// TIA Portal project "CLU" (V13)

(* hardware
DEVICE "S7-1200 station_1"  S7-1200 Station
   slot 0: "Telaio di montaggio_0"  Rack  V1.0
   slot 1: "S7_1200"  CPU 1214C DC/DC/DC  6ES7 214-1AG40-0XB0  V4.1
   slot 2: "DI 8/DQ 8x24VDC_1"  6ES7 223-1BH32-0XB0  V2.0
   slot 3: "DI 16/DQ 16x24VDC_1"  6ES7 223-1BL32-0XB0  V2.0
   slot 3: "Scheda di batteria_1"  6ES7 297-0AX30-0XA0  V1.0
   slot 4: "AI 8x13BIT_1"  6ES7 231-4HF32-0XB0  V2.0
   slot 5: "AI 8x13BIT_2"  6ES7 231-4HF32-0XB0  V2.0
   slot 6: "AQ 4x14BIT_1"  6ES7 232-4HD32-0XB0  V2.0
   slot 101: "CM 1241 (RS422/485)_1"  6ES7 241-1CH32-0XB0  V2.0
DEVICE "DISPLAY_KTP400"  KTP400 Basic color PN
   slot 0: "HMI"  HMI  6AV6 647-0AK11-3AX0  12.0.0.0
   slot 1: "HMI_RT_1"  KTP400 Basic color PN  6AV6 647-0AK11-3AX0  12.0.0.0
   slot 5: "DISPLAY_KTP400.IE_CP_1"  Interfaccia PROFINET
      slot 1: "PROFINET Interface_1"  Interfaccia PROFINET
         slot 1: "Porta_2"  Porta
*)

// ===== PLC "S7_1200"  CPU 1214C DC/DC/DC =====

VAR_GLOBAL   // PLC tag table "Tabella delle variabili standard"
   "ATTIVA_PRG" AT %M2.0 : Bool;   // Attiva il programma principale
   "System_Byte" AT %MB0 : Byte;
   "FirstScan" AT %M0.0 : Bool;   // Contatto chiuso solo alla prima scansiona
   "DiagStatusUpdate" AT %M0.1 : Bool;
   "AlwaysTRUE" AT %M0.2 : Bool;   // Contatto sempre chiuso
   "AlwaysFALSE" AT %M0.3 : Bool;   // Contatto sempre aperto
   "Clock_1.25Hz" AT %M1.4 : Bool;
   "Clock_1Hz" AT %M1.5 : Bool;
   "Clock_0.625Hz" AT %M1.6 : Bool;
   "Clock_0.5Hz" AT %M1.7 : Bool;
   "tasto_REMOTO" AT %I0.1 : Bool;
   "tasto_OFF" AT %I0.2 : Bool;
   "tasto_ON" AT %I0.3 : Bool;
   "tasto_ANODICA" AT %I0.4 : Bool;
   "tasto_RESET" AT %I0.5 : Bool;
   "led_LOCALE" AT %Q0.0 : Bool;
   "led_REMOTO" AT %Q0.1 : Bool;
   "led_OFF" AT %Q0.2 : Bool;
   "led_ON" AT %Q0.3 : Bool;
   "led_ANODICA" AT %Q0.4 : Bool;
   "led_RESET" AT %Q0.5 : Bool;
   "in_FLUSSO_LQD_TUBO_SEGNALE" AT %I0.6 : Bool;
   "in_FLUSSO_LQD_SS_SEGNALE" AT %I0.7 : Bool;
   "in_MAX_TEMP_LQD_SS_OK" AT %I1.0 : Bool;
   "in_MIN_PRESSIONE_LQD_SS_OK" AT %I1.1 : Bool;
   "in_INTERLOCK_OK" AT %I1.3 : Bool;
   "in_FLUSSO_LQD_TUBO_OK" AT %I1.4 : Bool;
   "in_FLUSSO_LQD_SS_OK" AT %I1.5 : Bool;
   "in_MAX_IG2_OK" AT %I2.0 : Bool;
   "adc_FWD_TUBO" AT %IW5 : Word;
   "adc_RFL_TUBO" AT %IW7 : Word;
   "adc_TENSIONE_ANODICA" AT %IW21 : Word;
   "adc_CORRENTE_ANODICA" AT %IW23 : Word;
   "adc_TENSIONE_G1" AT %IW25 : Word;
   "adc_CORRENTE_G1" AT %IW27 : Word;
   "adc_TENSIONE_G2" AT %IW29 : Word;
   "adc_CORRENTE_G2" AT %IW31 : Word;
   "led_RIFLESSA" AT %Q0.6 : Bool;
   "led_TEMPERTURA" AT %Q0.7 : Bool;
   "led_COOLING" AT %Q1.0 : Bool;
   "led_PREALLAME" AT %Q1.1 : Bool;
   "led_REDUCED" AT %Q2.0 : Bool;
   "led_NOMINAL" AT %Q2.1 : Bool;
   "in_PRESSIONE_ARIA_CAVITA_OK" AT %I3.0 : Bool;
   "in_PRESSIONE_ARIA_FILAMENTO_OK" AT %I3.1 : Bool;
   "in_ALIMENTAZIONE_G1_OK" AT %I3.3 : Bool;
   "in_ALIMENTAZIONE_G2_OK" AT %I3.4 : Bool;
   "in_MAX_TEMP_LQD_TUBO_OK" AT %I3.5 : Bool;
   "in_MIN_PRESSIONE_LQD_TUBO_OK" AT %I3.6 : Bool;
   "in_SLAVE_PREALLARME" AT %I2.7 : Bool;   // Ingresso modalità Master/Slave
   "in_CONDUCIMETRO_OK" AT %I4.0 : Bool;
   "in_ALTA_TENSIONE_OK" AT %I4.1 : Bool;
   "in_MAX_TEMP_TRASF_AT_OK" AT %I4.2 : Bool;
   "in_MANCANZA_FASE_OK" AT %I4.4 : Bool;
   "in_IGNITRON_OK" AT %I4.5 : Bool;
   "in_MAX_IA_OK" AT %I4.6 : Bool;
   "in_VALVOLA_CAVITA_OK" AT %I4.7 : Bool;
   "out_ON_PREAMPLIFICATORE" AT %Q4.6 : Bool;
   "out_ON_DRIVER" AT %Q4.7 : Bool;
   "out_ON_CW" AT %Q2.2 : Bool;
   "out_VENTILAZIONE_CAVITA" AT %Q3.0 : Bool;
   "out_SLAVE_RESET" AT %Q3.1 : Bool;   // Uscita modalità Master/Slave
   "out_ALIMENTAZIONE_FILAMENTO" AT %Q3.2 : Bool;
   "out_PARZIALIZZATORE_FILAMENTO" AT %Q4.4 : Bool;
   "out_ALIMENTAZIONE_G1" AT %Q3.3 : Bool;
   "out_PARZIALIZZATORE_AT" AT %Q4.5 : Bool;
   "out_ALIMENTAZIONE_G2" AT %Q3.4 : Bool;
   "out_G2" AT %Q3.5 : Bool;
   "adc_CORRENTE_FILAMENTO" AT %IW33 : Word;
   "adc_ANALOGICA_7" AT %IW35 : Word;   // DISPONIBILE ANALOGICA
   "tasto_LOCALE" AT %I0.0 : Bool;
   "out_SLAVE_ON" AT %Q2.3 : Bool;   // Uscita modalità Master/Slave
   "in_COAX_POS_B" AT %I1.2 : Bool;
   "in_COAX_POS_A" AT %I2.1 : Bool;
   "in_SAFETY_MODULE_OK" AT %I4.3 : Bool;
   "out_COAX" AT %Q2.4 : Bool;   // Comando posizione Coassiale (S)=B, (R)=A
   "out_SLAVE_OFF" AT %Q2.5 : Bool;   // Uscita modalità Master/Slave
   "out_ON_AMP1" AT %Q3.6 : Bool;
   "out_ON_AMP2" AT %Q3.7 : Bool;
   "out_IGNITRON" AT %Q4.0 : Bool;
   "out_SLAVE_ALLARME" AT %Q4.2 : Bool;   // Uscita modalità Master/Slave
   "out_SLAVE_ANODICA_OFF" AT %Q4.1 : Bool;   // Uscita modalità Master/Slave
   "adc_TEMP_LQDin_SS" AT %IW11 : Word;
   "adc_TEMP_LQDout_SS" AT %IW13 : Word;
   "adc_TEMP_LQDout_Tubo" AT %IW15 : Word;
   "adc_TEMP_LQDin_Tubo" AT %IW17 : Word;
   "adc_FWD_SS" AT %IW9 : Word;
   "adc_RFL_SS" AT %IW19 : Word;
   "adc_ANALOGICA_1" AT %IW38 : Word;
   "adc_ANALOGICA_2" AT %IW40 : Word;
   "in_SLAVE_ON" AT %I2.2 : Bool;   // Ingresso modalità Master/Slave
   "in_SLAVE_OFF" AT %I2.3 : Bool;   // Ingresso modalità Master/Slave
   "in_SLAVE_ANODICA_ON" AT %I2.4 : Bool;   // Ingresso modalità Master/Slave
   "in_SLAVE_ANODICA_OFF" AT %I2.5 : Bool;   // Ingresso modalità Master/Slave
   "in_SLAVE_ALLARME" AT %I2.6 : Bool;   // Ingresso modalità Master/Slave
   "in_SELECT_MODE" AT %I3.2 : Bool;   // Ingresso modalità Master/Slave
   "out_SLAVE_ANODICA_ON" AT %Q2.6 : Bool;
   "out_SLAVE_PREALLARME" AT %Q4.3 : Bool;   // Uscita modalità Master/Slave
   "out_CW_PULSED_TRIGGER" AT %Q2.7 : Bool;
   "in_SLAVE_RESET" AT %I3.7 : Bool;   // Ingresso modalità Master/Slave
   "dac_out_VA" AT %QW5 : Word;   // Uscita analogica regolatore Tensione di anodica
   "dac_out_VG2" AT %QW7 : Word;   // Uscita analogica regolatore Tensione di anodica
   "dac_out_VG1" AT %QW9 : Word;   // Uscita analogica regolatore Tensione di anodica
   "dac_out_VF" AT %QW11 : Word;   // Uscita analogica regolatore Tensione di anodica
END_VAR

DATA_BLOCK "STATO"   // DB1
TITLE = STATO AMPLIFICATORE
{ S7_Optimized_Access := 'FALSE' }
AUTHOR : Dario
VERSION : 0.1
// Blocco dati dello stato generale dell'amplificatore.
   VAR RETAIN
      stato_LOCALE : Bool;
      stato_STANDBY : Bool;
      stato_ANODICA : Bool;
      stato_ALLARME : Bool;
      stato_BLOCCO : Bool;
      stato_MODO_PULSED : Bool;
      stato_MODO_CW : Bool;
      stato_SOLO_SS : Bool;
      stato_NORMALE : Bool;
      stato_MASTER : Bool;
      stato_SLAVE : Bool;
   END_VAR
   VAR
      stato_RFridotta : Bool;
      stato_RFnominale : Bool;
   END_VAR
   VAR RETAIN
      stato_sogliaROS_Tubo : Word;
      stato_sogliaROS400kW : Word;
      stato_sogliaROS_SS_Pulsed : Word;
      "stato sogliaROS_SS_CW" : Word;
      stato_AQNdelay : Word;
      stato_LimiterInputRF : Word;
      stato_sogliaRIDOTTA : Word;
   END_VAR
   VAR
      stato_sogliaNOMINALE : Word;
   END_VAR
   VAR RETAIN
      stato_RFtotaleParziale : Bool;
   END_VAR
   VAR
      stato_DISPLAY_1 : Word;
      stato_DISPLAY_2 : Word;
      stato_DISPLAY_3 : Word;
      stato_DISPLAY_4 : Word;
      stato_DISPLAY_5 : Word;
      stato_DISPLAY_6 : Word;
   END_VAR
   VAR RETAIN
      stato_AdjFWDTubo : Word;
      stato_AdjRFLTubo : Word;
      stato_AdjFWDSS : Word;
      stato_AdjRFLSS : Word;
      stato_AdjFWDTotale : Word;
      stato_AdjRFLTotale : Word;
   END_VAR
   VAR
      stato_Data : DTL;
   END_VAR
   VAR RETAIN
      stato_ADDR_1 : Byte;
      stato_ADDR_2 : Byte;
      stato_ADDR_3 : Byte;
      stato_ADDR_4 : Byte;
      stato_PORT : UInt;
      stato_ADJ_ANODICA_PULSED : Word;
      stato_ADJ_ANODICA_CW : Word;
      stato_VOLTAGGIO_G1 : DInt;
      stato_VOLTAGGIO_G2 : Word;
      stato_VOLTAGGIO_FILAMENTO : Word;
      stato_REGOLAZIONE_VG1 : Word;
      stato_adj_VA : Word;
      stato_adj_VG1 : Word;
      stato_adj_VG2 : Word;
      stato_adj_VF : Word;
      stato_ScaleVA : Word;
      stato_ScaleVG1 : Word;
      stato_ScaleVG2 : Word;
      stato_ScaleIF : Word;
      stato_ScaleIA : Word;
      stato_ScaleIG1 : Word;
      stato_ScaleIG2 : Word;
   END_VAR
   VAR
      allarme_FLUSSO_LQD_TUBO : Bool;
      allarme_FLUSSO_LQD_SS : Bool;
      allarme_PRESSIONE_MIN_LQD_TUBO : Bool;
      allarme_PRESSIONE_MAX_LQD_TUBO : Bool;
      allarme_PRESSIONE_LQD_SS : Bool;
      allarme_INTERLOCK_RF : Bool;
      allarme_INTERLOCK_GENERALE : Bool;
      allarme_CONDUCIMETRO : Bool;
      allarme_MAX_IA : Bool;
      allarme_MAX_IG1 : Bool;
      allarme_MAX_IG2 : Bool;
      allarme_MAX_IG2_SW : Bool;
      allarme_TEMPERATURA_LQD_TUBO : Bool;
      allarme_TEMPERATURA_LQD_SS : Bool;
      allarme_TEMPERATURA_LQD_DUMMY : Bool;
      allarme_TEMPERATURA_AT : Bool;
      allarme_IGNITRON : Bool;
      allarme_ROS_Tubo : Bool;
      allarme_ROS_SS : Bool;
      allarme_No_Aria_Cavità : Bool;
      allarme_ROS_400kW : Bool;
      allarme_Assenza_VG1 : Bool;
      allarme_Assenza_VG2 : Bool;
      allarme_Assenza_AT : Bool;
      allarme_AMP1 : Bool;
      allarme_AMP2 : Bool;
      allarme_DRV : Bool;
      allarme_AMPcw : Bool;
      allarme_FASE : Bool;
      allarme_COAX : Bool;
      allarme_SAFETY : Bool;
      allarme_FILAMENTO : Bool;
      allarme_ANODICA_CW : Bool;
      allarme_SLAVE : Bool;
      allarme_MASTER : Bool;
      misura_TENSIONE_FILAMENTO : Word;
      misura_CORRENTE_FILAMENTO : Word;
      misura_TENSIONE_ANODICA : Word;
      misura_CORRENTE_ANODICA : Word;
      misura_TENSIONE_VG1 : Word;
      misura_CORRENTE_IG1 : Word;
      misura_TENSIONE_VG2 : Word;
      misura_CORRENTE_IG2 : Word;
      misura_FWD_Totale : Word;
      misura_RFL_Totale : Word;
      misura_FWD_TUBO : Word;
      misura_RFL_TUBO : Word;
      misura_FWD_SS : Word;
      misura_RFL_SS : Word;
      misura_TLQD_SS_Tin : Word;
      misura_TLQD_SS_Tout : Word;
      misura_FLQD_SS : Word;
      misura_TLQD_TUBO_Tin : Word;
      misura_TLQD_TUBO_Tout : Word;
      misura_FLQD_TUBO : Word;
   END_VAR
   VAR RETAIN
      misura_N_crowbar : Word;
   END_VAR
   VAR
      timer_Accensione_G1 : Word;
      timer_Spegnimento_G1 : Word;
      timer_PostVentilazione : Word;
      timer_AltaTensione : Word;
      timer_Accensione_G2 : Word;
      timer_Spegnimento_G2 : Word;
      timer_AccensioneSS : Word;
      controllo_ProcAccensione : Bool;
      controllo_ProcSpegnimento : Bool;
      controllo_AnodicaPronta : Bool;
      controllo_ProcAnodicaAccensione : Bool;
      controllo_ProcAnodicaSpegnimento : Bool;
      controllo_ProcSSAccensione : Bool;
      controllo_SpegnimentoPronto : Bool;
      controllo_ProcDriverAccensione : Bool;
      controllo_ImpostaOra : Bool;
      controllo_ProcReset : Bool;
      controllo_SetCModoCW : Bool;
      controllo_SetCModoIMPULSIVO : Bool;
      controllo_SetNormal : Bool;
      controllo_SetMaster : Bool;
      controllo_SetSlave : Bool;
      controllo_SetEPICS_IP : Bool;
      controllo_SetEPICS_Port : Bool;
      controllo_ResetSlave : Bool;
      controllo_SetParzialRF : Bool;
      controllo_SetTotalRF : Bool;
      controllo_ResetMaster : Bool;
      controllo_IgnoraSlave : Bool;
      controllo_changeAN_pulsed : Bool;
      controllo_changeAN_cw : Bool;
      controllo_setIG1Thr : Bool;
      controllo_setIG2Thr : Bool;
      controllo_setIFThr : Bool;
      controllo_setVG2 : Bool;
      controllo_setVG1 : Bool;
      controllo_setVF : Bool;
      controllo_ON_G1 : Bool;
      controllo_setReduced : Bool;
      controllo_EnEPICS : Bool;
      tlc_ampli_ON : Bool;
      tlc_ampli_OFF : Bool;
      tlc_ampli_ANODICA_ON : Bool;
      tlc_ampli_ANODICA_OFF : Bool;
      tlc_ampli_RESET : Bool;
      tlc_set_NORMAL : Bool;
      tlc_set_MASTER : Bool;
      tlc_set_SLAVE : Bool;
      tlc_enable_400kW : Bool;
      tlc_disable_400kW : Bool;
      tlc_set_DAC_Anodica : Bool;
      tlc_set_IG1 : Bool;
      tlc_set_IG2 : Bool;
      tlc_set_IF : Bool;
      tlc_set_VG1 : Bool;
      tlc_set_VG2 : Bool;
      tlc_set_VF : Bool;
      tlc_Dac_value : Word;
      tlc_IG1_value : Word;
      tlc_IG2_value : Word;
      tlc_IF_value : Word;
      tlc_VG1_value : Word;
      tlc_VG2_value : Word;
      tlc_VF_value : Word;
   END_VAR
   VAR RETAIN
      TIMEOUT_preheating : Int;
      TIMEOUT_cooldown : Int;
      TIMEOUT_postVentilazione : Int;
      TIMEOUT_initAT : Int;
      TIMEOUT_initG2 : Int;
      TIMEOUT_initSS : Int;
      TIMEOUT_stopG2 : Int;
      SOGLIA_IFonG1 : Int;
      SOGLIA_VAcw : Int;
      SOGLIA_IG1 : Int;
      SOGLIA_IG2 : Int;
      info_SW_revisione : Int;
   END_VAR
   VAR
      SIGNED_G1_VOLTAGE : DInt;
   END_VAR
   VAR RETAIN
      divisore_TUBO : Int;
   END_VAR
   VAR
      FWD_DISPLAY : Word;
      RFL_DISPLAY : Word;
      FWD_DISPLAY_BARRA : Word;
      RFL_DISPLAY_BARRA : Word;
   END_VAR
   VAR RETAIN
      MAX_THR_RFL_TUBO : Word;
   END_VAR
   VAR
      valore : Int;
   END_VAR
   VAR RETAIN
      SogliaRidotta : Word;
      adj_Tube_CW_FWD : Word;
      adj_Tube_CW_RFL : Word;
   END_VAR
BEGIN
END_DATA_BLOCK

DATA_BLOCK "MAIN_PRG_DB"   // DB4
{ S7_Optimized_Access := 'FALSE' }
VERSION : 0.1
// stored: InstanceOfName MAIN_PRG
"MAIN_PRG"
BEGIN
END_DATA_BLOCK

DATA_BLOCK "STATO_TMP"   // DB7
{ S7_Optimized_Access := 'FALSE' }
VERSION : 0.1
   VAR
      tmp_flussoTubo_LQD : Word;
      tmp_flussoSS_LQD : Word;
      tmp_timer_flussoTubo : Word;
      tmp_timer_flussoSS : Word;
      tmp_Data : DTL;
      tmp_setDelay : Bool;
      tmp_setLimiter : Bool;
      tmp_sogliaRFnominale : DInt;
      tmp_adj_anodica_pulsed : Word;
      tmp_adj_anodica_cw : Word;
      tmp_adj_VG2 : Word;
      tmp_IG1 : Word;
      tmp_IG2 : Word;
      tmp_IF : Word;
      tmp_Reduced : Word;
      tmp_real_VG2 : Real;
      tmp_real_Anodica : Real;
      tmp_adj_VA : DInt;
      tmp_adj_VG1 : DInt;
      tmp_adj_G1 : DInt;
      tmp_adj_G2 : DInt;
      tmp_adj_VF : DInt;
      tmp_VG1r : Real;
      tmp_VFr : Real;
      tmpVFi : Word;
      tmp_VFin : Word;
      tmp_VFctrl : Bool;
      tmp_timerG1 : Word;
      tmp_error : Bool;
      tmp_errorCode : Word;
   END_VAR
BEGIN
END_DATA_BLOCK

DATA_BLOCK "TABELLE_LINEARIZZAZIONE"   // DB12
{ S7_Optimized_Access := 'FALSE' }
VERSION : 0.1
   VAR
      tab_TUBO_Pulsed : Array[0..32] of Word;
      tab_TUBO_CW : Array[0..32] of Word;
      tab_SS_Pulsed : Array[0..32] of Word;
      tab_SS_CW : Array[0..32] of Word;
      tab_TOTALE : Array[0..32] of Word;
      tab_TOTALE_CW : Array[0..32] of Word;
      tab_Vanodica : Array[0..36] of Word;
      tab_VG1 : Array[0..14] of Int;
   END_VAR
BEGIN
END_DATA_BLOCK

DATA_BLOCK "SERIAL_DATA"   // DB15
{ S7_Optimized_Access := 'FALSE' }
VERSION : 0.1
   VAR
      messaggio_76h : Array[0..4] of Byte;
      mesaggio_46h : Array[0..8] of Byte;
      messaggio_49h : Array[0..11] of Byte;
      buffer_ricezione : Array[0..99] of Byte;
      trasmissioneAbilitata : Bool;
      AttivoInvio : Bool;
      FermaInvio : Bool;
      CominciaRicezione : Bool;
      RS485doneTX : Bool;
      RS485errorTX : Bool;
      RS485doneRX : Bool;
      RS485errorRX : Bool;
      RS485statusTX : Word;
      RS485statusRX : Word;
      comandoInCoda : Word;
      ADDRESS : Word;
      ADDR_RCV : Word;
      NEXT_SLAVE : Word;
      BYTE_RICEVUTI : Word;
      faultContatoreAMP1 : Word;
      faultContatoreAMP2 : Word;
      faultContatoreDRV : Word;
      faultContatoreAMPcw : Word;
      LRC_messaggio : Byte;
      LRC_calcolato : Byte;
   END_VAR
BEGIN
END_DATA_BLOCK

DATA_BLOCK "SLAVE_DATA"   // DB21
TITLE = SLAVE_DATA
{ S7_Optimized_Access := 'FALSE' }
AUTHOR : Dario
VERSION : 0.1
// Blocco dati che contiene i parametri letti dalla RS2485 degli amplificatori dello Stato Solido, più le scheda Delay e RF Limiter.
   VAR
      AMP1_Allarmi : Word;
      AMP1_V1 : Word;
      AMP1_V2 : Word;
      AMP1_I1 : Word;
      AMP1_I2 : Word;
      AMP1_I3 : Word;
      AMP1_I4 : Word;
      AMP1_I5 : Word;
      AMP1_I6 : Word;
      AMP1_I7 : Word;
      AMP1_I8 : Word;
      AMP1_FWD : Word;
      AMP1_RFL : Word;
      AMP1_IN : Word;
      AMP1_TMP : Word;
      AMP2_Allarmi : Word;
      AMP2_V1 : Word;
      AMP2_V2 : Word;
      AMP2_I1 : Word;
      AMP2_I2 : Word;
      AMP2_I3 : Word;
      AMP2_I4 : Word;
      AMP2_I5 : Word;
      AMP2_I6 : Word;
      AMP2_I7 : Word;
      AMP2_I8 : Word;
      AMP2_FWD : Word;
      AMP2_RFL : Word;
      AMP2_IN : Word;
      AMP2_TMP : Word;
      DRV_Allarmi : Word;
      DRV_V1 : Word;
      DRV_I1 : Word;
      DRV_FWD : Word;
      DRV_RFL : Word;
      DRV_TMP : Word;
      AMPcw_Allarmi : Word;
      AMPcw_Vd : Word;
      AMPcw_V1 : Word;
      AMPcw_V2 : Word;
      AMPcw_Id : Word;
      AMPcw_I1 : Word;
      AMPcw_I2 : Word;
      AMPcw_FWD : Word;
      AMPcw_RFL : Word;
      AMPcw_IN : Word;
      AMPcw_TMP : Word;
      AQN_Allarmi : Word;
      AQN_Delay : Word;
      LIM_Allarmi : Word;
      LIM_value : Word;
   END_VAR
BEGIN
END_DATA_BLOCK

DATA_BLOCK "EPICS_READ"   // DB27
{ S7_Optimized_Access := 'FALSE' }
VERSION : 0.1
   VAR
      STATO_LOCALE : Word;
      STATO_STANDBY : Word;
      STATO_ANODICA : Word;
      STATO_ALLARME : Word;
      STATO_FAULT : Word;
      STATO_MODO_IC : Word;
      STATO_MODO_MS : Word;
      MIN_PRESSIONE_ARIA_CAVITA : Word;
      MAX_REFL_400KW : Word;
      MIN_FLUSSO_LQD_TUBO : Word;
      MIN_PRESSIONE_LQD_TUBO : Word;
      MAX_TEMP_LQD_TUBO : Word;
      MIN_FLUSSO_LQD_SS : Word;
      MIN_PRESSIONE_LQD_SS : Word;
      MAX_TEMP_LQD_SS : Word;
      INTERLOCK_OPEN : Word;
      IA_MAX : Word;
      IG1_MAX : Word;
      IG2_MAX : Word;
      INTERVENTO_SCR : Word;
      PHASE_FAIL : Word;
      NO_VG1 : Word;
      NO_VG2 : Word;
      MAX_REFL_TUBO : Word;
      MAX_REFL_SS : Word;
      MISURA_TENSIONE_FILAMENTO : Word;
      MISURA_CORRENTE_FILAMENTO : Word;
      MISURA_TENSIONE_G1 : Word;
      MISURA_CORRENTE_G1 : Word;
      MISURA_TENSIONE_G2 : Word;
      MISURA_CORRENTE_G2 : Word;
      MISURA_TENSIONE_ANODICA : Word;
      MISURA_CORRENTE_ANODICA : Word;
      MISURA_FWD_TUBO : Word;
      MISURA_REFL_TUBO : Word;
      MISURA_FWD_SS : Word;
      MISURA_REFL_SS : Word;
      MISURA_FLUSSO_LQD_TUBO : Word;
      MISURA_FLUSSO_LQD_SS : Word;
      MISURA_TEMPERATURA_LQD_IN_TUBO : Word;
      MISURA_TEMPERATURA_LQD_OUT_TUBO : Word;
      MISURA_TEMPERATURA_LQD_IN_SS : Word;
      MISURA_TEMPERATURA_LQD_OUT_SS : Word;
      TEMPO_RISCALDAMENTO_FILAMENTO : Word;
      TEMPO_COOLDOWN_FILAMENTO : Word;
      TEMPO_POSTVENTILAZIONE : Word;
      AMPLI1_V1 : Word;
      AMPLI1_V2 : Word;
      AMPLI1_I1 : Word;
      AMPLI1_I2 : Word;
      AMPLI1_I3 : Word;
      AMPLI1_I4 : Word;
      AMPLI1_I5 : Word;
      AMPLI1_I6 : Word;
      AMPLI1_I7 : Word;
      AMPLI1_I8 : Word;
      AMPLI1_FWD : Word;
      AMPLI1_RFL : Word;
      AMPLI1_TMP : Word;
      AMPLI2_V1 : Word;
      AMPLI2_V2 : Word;
      AMPLI2_I1 : Word;
      AMPLI2_I2 : Word;
      AMPLI2_I3 : Word;
      AMPLI2_I4 : Word;
      AMPLI2_I5 : Word;
      AMPLI2_I6 : Word;
      AMPLI2_I7 : Word;
      AMPLI2_I8 : Word;
      AMPLI2_FWD : Word;
      AMPLI2_RFL : Word;
      AMPLI2_TMP : Word;
      DRV_V1 : Word;
      DRV_I1 : Word;
      DRV_FWD : Word;
      DRV_RFL : Word;
      DRV_TMP : Word;
      AMPLIcw_VD : Word;
      AMPLIcw_V1 : Word;
      AMPLIcw_V2 : Word;
      AMPLIcw_ID : Word;
      AMPLIcw_I1 : Word;
      AMPLIcw_I2 : Word;
      AMPLIcw_FWD : Word;
      AMPLIcw_RFL : Word;
      AMPLIcw_TMP : Word;
      STATE_400_SAMPLING : Word;
      N_CROWBAR : Word;
      FWD_TOTAL : Word;
      RFL_TOTAL : Word;
      DAC_ANODICA_PULSED : Word;
      DAC_ANODICA_CW : Word;
      SOGLIA_IG1 : Word;
      SOGLIA_IG2 : Word;
      SOGLIA_IF : Word;
      ALM_SAFETY : Word;
      ALM_FILAMENT : Word;
      ALM_CW_ANODICA : Word;
      ALM_ALTA_TENSIONE : Word;
      ALM_TEMP_ALTA_TENSIONE : Word;
      ALM_CONDUCIMETER : Word;
      ALM_COAX : Word;
      ALM_SLAVE : Word;
      ALM_MASTER : Word;
      REGOLAZIONE_VG1 : Word;
      REGOLAZIONE_VG2 : Word;
      REGOLAZIONE_VF : Word;
      TLS_FREE_1 : Word;
      TLS_FREE_2 : Word;
      TLS_FREE_3 : Word;
   END_VAR
BEGIN
END_DATA_BLOCK

DATA_BLOCK "EPICS_WRITE"   // DB28
{ S7_Optimized_Access := 'FALSE' }
VERSION : 0.1
   VAR
      TLC_ON : Word;
      TLC_OFF : Word;
      TLC_ANODICA_ON : Word;
      TLC_ANODICA_OFF : Word;
      TLC_RESET : Word;
      TLC_SET_NORMAL : Word;
      TLC_SET_MASTER : Word;
      TLC_SET_SLAVE : Word;
      TLC_ENABLE_400kW : Word;
      TLC_DISABLE_400kW : Word;
      TLC_ANODIC_PULSED_VOLTAGE : Word;
      TLC_ANODIC_CW_VOLTAGE : Word;
      TLC_IG1_MAX_THR : Word;
      TLC_IG2_MAX_THR : Word;
      TLC_IF_MIN_THR : Word;
      TLC_SET_VA : Word;
      TLC_SET_IG1 : Word;
      TLC_SET_IG2 : Word;
      TLC_SET_IF : Word;
      TLC_VG1_VALUE : Word;
      TLC_VG2_VALUE : Word;
      TLC_VF_VALUE : Word;
      TLC_SET_VG1 : Word;
      TLC_SET_VG2 : Word;
      TLC_SET_VF : Word;
      TLC_FREE_1 : Word;
      TLC_FREE_2 : Word;
      TLC_FREE_3 : Word;
   END_VAR
BEGIN
END_DATA_BLOCK

DATA_BLOCK "ETHERNET_CTRL"   // DB29
{ S7_Optimized_Access := 'FALSE' }
VERSION : 0.1
   VAR
      START_eth_SEND : Bool;
      START_eth_RECV : Bool;
      STATO_TX_Connection : Bool;
      STATO_RX_Connection : Bool;
      Restart_Block_TX : Bool;
      Restart_Block_RX : Bool;
      TCP_CONN_DONE : Bool;
      TCP_TX_DONE : Bool;
      TCP_RX_DONE : Bool;
      TCP_CONN_BUSY : Bool;
      TCP_TX_BUSY : Bool;
      TCP_RX_BUSY : Bool;
      TCP_CONN_ERROR : Bool;
      TCP_TX_ERROR : Bool;
      TCP_RX_ERROR : Bool;
      TCP_CONN_STATUS : Word;
      TCP_TX_STATUS : Word;
      TCP_RX_STATUS : Word;
      N_RECEIVED_DATA : Word;
   END_VAR
BEGIN
END_DATA_BLOCK

// folder: System blocks/Program resources

DATA_BLOCK "IEC_Timer_0_DB"   // DB3
{ S7_Optimized_Access := 'FALSE' }
AUTHOR : Simatic
FAMILY : IEC
NAME : IEC_TMR
VERSION : 1.0
// stored: InstanceOfName ?
"?"
BEGIN
END_DATA_BLOCK

DATA_BLOCK "Timeout_AMP"   // DB5
{ S7_Optimized_Access := 'FALSE' }
AUTHOR : Simatic
FAMILY : IEC
NAME : IEC_TMR
VERSION : 1.0
// stored: InstanceOfName ?
"?"
BEGIN
END_DATA_BLOCK

DATA_BLOCK "Timeout_DRV"   // DB6
{ S7_Optimized_Access := 'FALSE' }
AUTHOR : Simatic
FAMILY : IEC
NAME : IEC_TMR
VERSION : 1.0
// stored: InstanceOfName ?
"?"
BEGIN
END_DATA_BLOCK

DATA_BLOCK "Timeout_AT"   // DB8
{ S7_Optimized_Access := 'FALSE' }
AUTHOR : Simatic
FAMILY : IEC
NAME : IEC_TMR
VERSION : 1.0
// stored: InstanceOfName ?
"?"
BEGIN
END_DATA_BLOCK

DATA_BLOCK "Timeout_VG1"   // DB9
{ S7_Optimized_Access := 'FALSE' }
AUTHOR : Simatic
FAMILY : IEC
NAME : IEC_TMR
VERSION : 1.0
// stored: InstanceOfName ?
"?"
BEGIN
END_DATA_BLOCK

DATA_BLOCK "Timeout_SorgenteRF"   // DB10
{ S7_Optimized_Access := 'FALSE' }
AUTHOR : Simatic
FAMILY : IEC
NAME : IEC_TMR
VERSION : 1.0
// stored: InstanceOfName ?
"?"
BEGIN
END_DATA_BLOCK

DATA_BLOCK "Timeout_VG2"   // DB11
{ S7_Optimized_Access := 'FALSE' }
AUTHOR : Simatic
FAMILY : IEC
NAME : IEC_TMR
VERSION : 1.0
// stored: InstanceOfName ?
"?"
BEGIN
END_DATA_BLOCK

DATA_BLOCK "Timeout_Ventilazione_Cavità"   // DB13
{ S7_Optimized_Access := 'FALSE' }
AUTHOR : Simatic
FAMILY : IEC
NAME : IEC_TMR
VERSION : 1.0
// stored: InstanceOfName ?
"?"
BEGIN
END_DATA_BLOCK

DATA_BLOCK "timeout_reset_ETH"   // DB14
{ S7_Optimized_Access := 'FALSE' }
AUTHOR : Simatic
FAMILY : IEC
NAME : IEC_TMR
VERSION : 1.0
// stored: InstanceOfName ?
"?"
BEGIN
END_DATA_BLOCK

DATA_BLOCK "Timeout_RS485_TX"   // DB16
{ S7_Optimized_Access := 'FALSE' }
AUTHOR : Simatic
FAMILY : IEC
NAME : IEC_TMR
VERSION : 1.0
// stored: InstanceOfName ?
"?"
BEGIN
END_DATA_BLOCK

DATA_BLOCK "Timeout_CambioAQN"   // DB22
{ S7_Optimized_Access := 'FALSE' }
AUTHOR : Simatic
FAMILY : IEC
NAME : IEC_TMR
VERSION : 1.0
// stored: InstanceOfName ?
"?"
BEGIN
END_DATA_BLOCK

DATA_BLOCK "Timeout_CambioLimiter"   // DB23
{ S7_Optimized_Access := 'FALSE' }
AUTHOR : Simatic
FAMILY : IEC
NAME : IEC_TMR
VERSION : 1.0
// stored: InstanceOfName ?
"?"
BEGIN
END_DATA_BLOCK

DATA_BLOCK "Timeout_NominaleVeloce"   // DB24
{ S7_Optimized_Access := 'FALSE' }
AUTHOR : Simatic
FAMILY : IEC
NAME : IEC_TMR
VERSION : 1.0
// stored: InstanceOfName ?
"?"
BEGIN
END_DATA_BLOCK

DATA_BLOCK "Timeout_NominaleLento"   // DB25
{ S7_Optimized_Access := 'FALSE' }
AUTHOR : Simatic
FAMILY : IEC
NAME : IEC_TMR
VERSION : 1.0
// stored: InstanceOfName ?
"?"
BEGIN
END_DATA_BLOCK

DATA_BLOCK "Timeout_Coassiale"   // DB26
{ S7_Optimized_Access := 'FALSE' }
AUTHOR : Simatic
FAMILY : IEC
NAME : IEC_TMR
VERSION : 1.0
// stored: InstanceOfName ?
"?"
BEGIN
END_DATA_BLOCK

DATA_BLOCK "Timeout_ETH_Send"   // DB30
{ S7_Optimized_Access := 'FALSE' }
AUTHOR : Simatic
FAMILY : IEC
NAME : IEC_TMR
VERSION : 1.0
// stored: InstanceOfName ?
"?"
BEGIN
END_DATA_BLOCK

DATA_BLOCK "S7_1200_Send_DB"   // DB32
{ S7_Optimized_Access := 'FALSE' }
AUTHOR : SIMATIC
FAMILY : MC7Plus
NAME : TC_IP_v4
VERSION : 1.0
// stored: InstanceOfName ?
"?"
BEGIN
END_DATA_BLOCK

DATA_BLOCK "Timeout_Ripristino_TX"   // DB33
{ S7_Optimized_Access := 'FALSE' }
AUTHOR : Simatic
FAMILY : IEC
NAME : IEC_TMR
VERSION : 1.0
// stored: InstanceOfName ?
"?"
BEGIN
END_DATA_BLOCK

DATA_BLOCK "Timeout_ETH_Recv"   // DB34
{ S7_Optimized_Access := 'FALSE' }
AUTHOR : Simatic
FAMILY : IEC
NAME : IEC_TMR
VERSION : 1.0
// stored: InstanceOfName ?
"?"
BEGIN
END_DATA_BLOCK

DATA_BLOCK "Timeout_Ripristino_RX"   // DB36
{ S7_Optimized_Access := 'FALSE' }
AUTHOR : Simatic
FAMILY : IEC
NAME : IEC_TMR
VERSION : 1.0
// stored: InstanceOfName ?
"?"
BEGIN
END_DATA_BLOCK

DATA_BLOCK "IEC_Timer_0_DB_1"   // DB45
{ S7_Optimized_Access := 'FALSE' }
AUTHOR : Simatic
FAMILY : IEC
NAME : IEC_TMR
VERSION : 1.0
// stored: InstanceOfName ?
"?"
BEGIN
END_DATA_BLOCK

DATA_BLOCK "IEC_Timer_0_DB_2"   // DB46
{ S7_Optimized_Access := 'FALSE' }
AUTHOR : Simatic
FAMILY : IEC
NAME : IEC_TMR
VERSION : 1.0
// stored: InstanceOfName ?
"?"
BEGIN
END_DATA_BLOCK

DATA_BLOCK "timeout_Max_IG1"   // DB47
{ S7_Optimized_Access := 'FALSE' }
AUTHOR : Simatic
FAMILY : IEC
NAME : IEC_TMR
VERSION : 1.0
// stored: InstanceOfName ?
"?"
BEGIN
END_DATA_BLOCK

DATA_BLOCK "timeout_Enable_G2"   // DB48
{ S7_Optimized_Access := 'FALSE' }
AUTHOR : Simatic
FAMILY : IEC
NAME : IEC_TMR
VERSION : 1.0
// stored: InstanceOfName ?
"?"
BEGIN
END_DATA_BLOCK

DATA_BLOCK "timeout_FLOW_SS"   // DB49
{ S7_Optimized_Access := 'FALSE' }
AUTHOR : Simatic
FAMILY : IEC
NAME : IEC_TMR
VERSION : 1.0
// stored: InstanceOfName ?
"?"
BEGIN
END_DATA_BLOCK

DATA_BLOCK "timeout_FLOW_TUBE"   // DB50
{ S7_Optimized_Access := 'FALSE' }
AUTHOR : Simatic
FAMILY : IEC
NAME : IEC_TMR
VERSION : 1.0
// stored: InstanceOfName ?
"?"
BEGIN
END_DATA_BLOCK

DATA_BLOCK "timeout_init_AT"   // DB51
{ S7_Optimized_Access := 'FALSE' }
AUTHOR : Simatic
FAMILY : IEC
NAME : IEC_TMR
VERSION : 1.0
// stored: InstanceOfName ?
"?"
BEGIN
END_DATA_BLOCK

DATA_BLOCK "timeout_stop_G1"   // DB52
{ S7_Optimized_Access := 'FALSE' }
AUTHOR : Simatic
FAMILY : IEC
NAME : IEC_TMR
VERSION : 1.0
// stored: InstanceOfName ?
"?"
BEGIN
END_DATA_BLOCK

DATA_BLOCK "timerChangeVF"   // DB54
{ S7_Optimized_Access := 'FALSE' }
AUTHOR : Simatic
FAMILY : IEC
NAME : IEC_TMR
VERSION : 1.0
// stored: InstanceOfName ?
"?"
BEGIN
END_DATA_BLOCK

// folder: (top level)

FUNCTION_BLOCK "MAIN_PRG"   // FB1, LAD
TITLE = PROGRAMMA PRINCIPALE
{ S7_Optimized_Access := 'FALSE' }
VERSION : 0.1
   VAR_TEMP   // added for the SCL form of the ladder/FBD networks
      _w1 : Bool;
      _w2 : Bool;
      _w3 : Bool;
      _w4 : Bool;
   END_VAR
BEGIN

REGION Network 1: Lettura orologio
   // Leggo la data corrente.
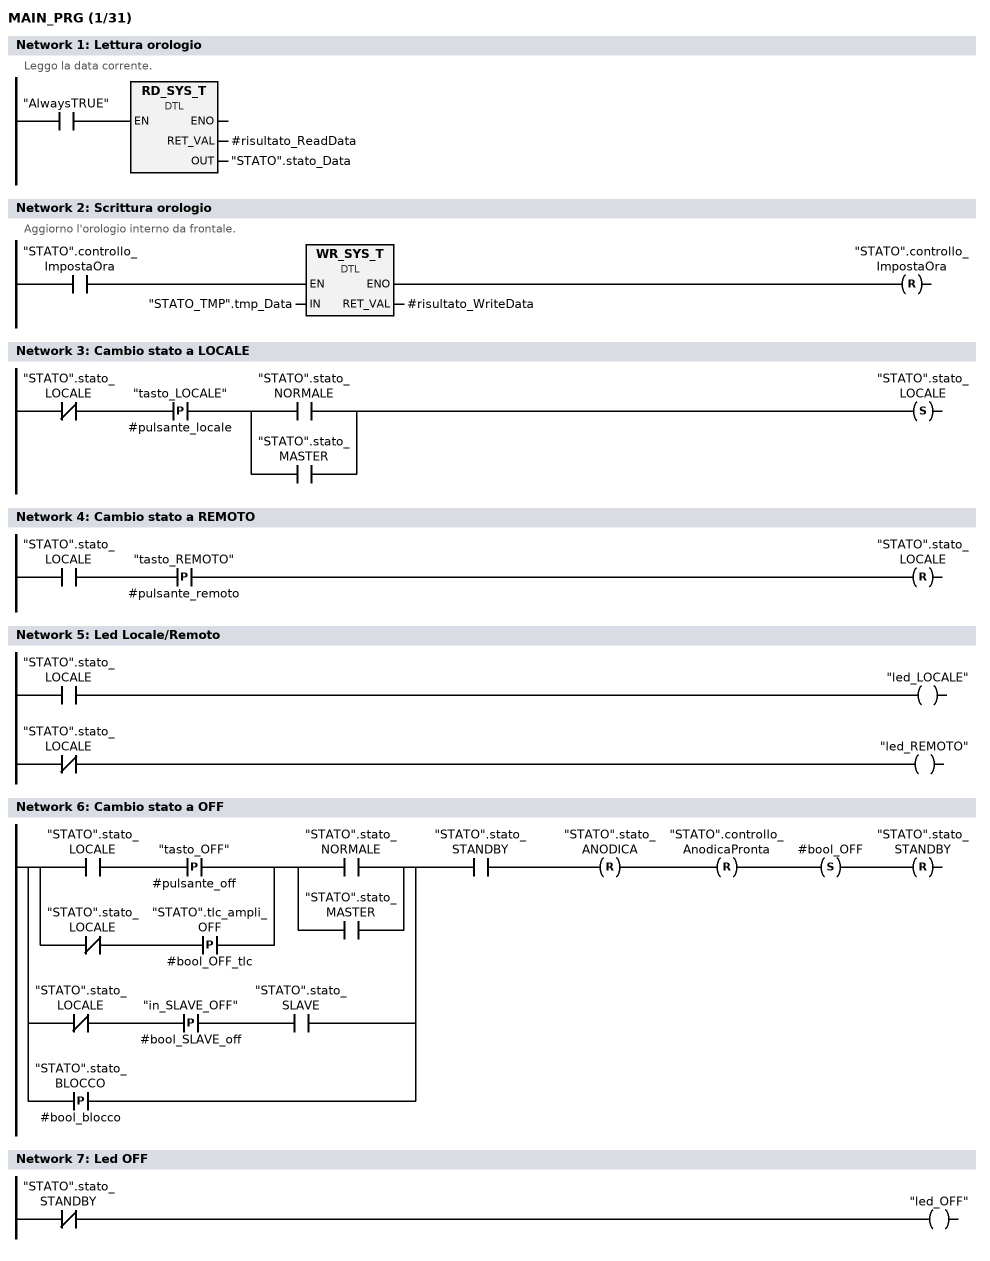
   IF "AlwaysTRUE" THEN #risultato_ReadData := RD_SYS_T(OUT => "STATO".stato_Data); END_IF;
END_REGION

REGION Network 2: Scrittura orologio
   // Aggiorno l'orologio interno da frontale.
   // ENO of a box is taken as its EN; it also drops when the box reports an error
   #_w1 := "STATO".controllo_ImpostaOra;
   IF #_w1 THEN
       #risultato_WriteData := WR_SYS_T(IN := "STATO_TMP".tmp_Data);
       "STATO".controllo_ImpostaOra := FALSE;
   END_IF;
END_REGION

REGION Network 3: Cambio stato a LOCALE
   RUNG wire#powerrail
      I_Contact( "STATO".stato_LOCALE )
      P_Contact(operand := "tasto_LOCALE", bit := #pulsante_locale)
      wire#w1
      Contact( "STATO".stato_NORMALE )
      wire#w2
      S_Coil( "STATO".stato_LOCALE )
   END_RUNG
   RUNG wire#w1
      Contact( "STATO".stato_MASTER )
   END_RUNG wire#w2
   // the same network as SCL:
   #_w1 := NOT "STATO".stato_LOCALE AND "tasto_LOCALE" AND NOT #pulsante_locale;   // rising edge of "tasto_LOCALE"
   #pulsante_locale := "tasto_LOCALE";
   IF #_w1 AND ("STATO".stato_NORMALE OR "STATO".stato_MASTER) THEN "STATO".stato_LOCALE := TRUE; END_IF;
END_REGION

REGION Network 4: Cambio stato a REMOTO
   RUNG wire#powerrail
      Contact( "STATO".stato_LOCALE )
      P_Contact(operand := "tasto_REMOTO", bit := #pulsante_remoto)
      R_Coil( "STATO".stato_LOCALE )
   END_RUNG
   // the same network as SCL:
   #_w1 := "STATO".stato_LOCALE AND "tasto_REMOTO" AND NOT #pulsante_remoto;   // rising edge of "tasto_REMOTO"
   #pulsante_remoto := "tasto_REMOTO";
   IF #_w1 THEN "STATO".stato_LOCALE := FALSE; END_IF;
END_REGION

REGION Network 5: Led Locale/Remoto
   RUNG wire#powerrail
      Contact( "STATO".stato_LOCALE )
      Coil( "led_LOCALE" )
   END_RUNG
   RUNG wire#powerrail
      I_Contact( "STATO".stato_LOCALE )
      Coil( "led_REMOTO" )
   END_RUNG
   // the same network as SCL:
   "led_LOCALE" := "STATO".stato_LOCALE;
   "led_REMOTO" := NOT "STATO".stato_LOCALE;
END_REGION

REGION Network 6: Cambio stato a OFF
   RUNG wire#powerrail
      Contact( "STATO".stato_LOCALE )
      P_Contact(operand := "tasto_OFF", bit := #pulsante_off)
      wire#w1
      Contact( "STATO".stato_NORMALE )
      wire#w2
      Contact( "STATO".stato_STANDBY )
      R_Coil( "STATO".stato_ANODICA )
      R_Coil( "STATO".controllo_AnodicaPronta )
      S_Coil( #bool_OFF )
      R_Coil( "STATO".stato_STANDBY )
   END_RUNG
   RUNG wire#powerrail
      I_Contact( "STATO".stato_LOCALE )
      P_Contact(operand := "STATO".tlc_ampli_OFF, bit := #bool_OFF_tlc)
   END_RUNG wire#w1
   RUNG wire#w1
      Contact( "STATO".stato_MASTER )
   END_RUNG wire#w2
   RUNG wire#powerrail
      I_Contact( "STATO".stato_LOCALE )
      P_Contact(operand := "in_SLAVE_OFF", bit := #bool_SLAVE_off)
      Contact( "STATO".stato_SLAVE )
   END_RUNG wire#w2
   RUNG wire#powerrail
      P_Contact(operand := "STATO".stato_BLOCCO, bit := #bool_blocco)
   END_RUNG wire#w2
   // the same network as SCL:
   #_w1 := "STATO".stato_LOCALE AND "tasto_OFF" AND NOT #pulsante_off;   // rising edge of "tasto_OFF"
   #pulsante_off := "tasto_OFF";
   #_w2 := NOT "STATO".stato_LOCALE AND "STATO".tlc_ampli_OFF AND NOT #bool_OFF_tlc;   // rising edge of "STATO".tlc_ampli_OFF
   #bool_OFF_tlc := "STATO".tlc_ampli_OFF;
   #_w3 := NOT "STATO".stato_LOCALE AND "in_SLAVE_OFF" AND NOT #bool_SLAVE_off;   // rising edge of "in_SLAVE_OFF"
   #bool_SLAVE_off := "in_SLAVE_OFF";
   #_w4 := "STATO".stato_BLOCCO AND NOT #bool_blocco;   // rising edge of "STATO".stato_BLOCCO
   #bool_blocco := "STATO".stato_BLOCCO;
   IF (((#_w1 OR #_w2) AND ("STATO".stato_NORMALE OR "STATO".stato_MASTER)) OR (#_w3 AND "STATO".stato_SLAVE) OR #_w4) AND "STATO".stato_STANDBY THEN
       "STATO".stato_ANODICA := FALSE;
       "STATO".controllo_AnodicaPronta := FALSE;
       #bool_OFF := TRUE;
       "STATO".stato_STANDBY := FALSE;
   END_IF;
END_REGION

REGION Network 7: Led OFF
   RUNG wire#powerrail
      I_Contact( "STATO".stato_STANDBY )
      Coil( "led_OFF" )
   END_RUNG
   // the same network as SCL:
   "led_OFF" := NOT "STATO".stato_STANDBY;
END_REGION

REGION Network 8: Cambio stato a ON
   // Se no allarmi passo in stato ON